(* Logix 5000 project; controller FV vendor 1 type 14 code 217 rev 31.11; software revision 31.00 *) (continued)
   FR_N10 : INT[265] := ([1] := 1, [2] := 4, [3] := 6, [6] := 6, [100] := 1, [101] := 2, [102] := 3, [103] := 3, [104] := 9, [105] := 9, [106] := 3, [200] := 2, [203] := 20, [204] := 191, [205] := 137, [206] := 100, [209] := 23, [215] := 14641, [216] := 11826, [217] := 13873, [218] := 11832, [219] := 12338, [220] := 13102, [221] := 49);   // FV_AGING Comms to FV Aging PL C
        [0]   // FV Unit Heartbeat
        [0].0   // FV_Aging PLC Heartbeat
        [100].0   // FV Routing (This)PLC Heartbeat
        [101]   // FV26 Routing Status to FV PLC
        [102]   // FV27 Routing Status to FV PLC
        [103]   // FV28 Routing Status to FV PLC
        [104]   // FV29 Routing Status to FV PLC
        [105]   // FV30 Routing Status to FV PLC
        [106]   // FV31 Routing Status to FV PLC
        [1]   // FV26 Aging Status from FV PLC
        [200].0   // FV_Aging_PLC Heartbeat Fault
        [200].1   // Enable Comms to FV Aging PLC
        [201]   // FV_Aging PLC Comms Control Block
        [2]   // FV27 Aging Status from FV PLC
        [3]   // FV28 Aging Status from FV PLC
        [4]   // FV29 Aging Status from FV PLC
        [5]   // FV30 Aging Status from FV PLC
        [6]   // FV31 Aging Status from FV PLC
   FR_N100 : INT[265] := ([2] := 1, [3] := 129, [6] := -1, [7] := -1, [8] := 2530, [9] := -1, [10] := 1, [15] := 1, [20] := -1, [21] := -1, [22] := -1, [23] := -1, [24] := -1, [25] := -1, [26] := -1, [30] := 226, [32] := 1000, [33] := 8, [35] := -1, [36] := -1, [40] := 26, [42] := 70, [47] := 50, [48] := 300, [49] := 32760, [57] := 2046, [70] := 32760, [71] := 32760, [72] := 32760, [73] := 32760, [74] := 32760, [75] := 32760, [100] := 22, [101] := 9, [102] := 14, [103] := 26, [104] := 25, [105] := 37, [106] := 28, [107] := 33, [108] := 41, [109] := 40, [110] := 74, [111] := 65, [112] := 70, [113] := 78, [114] := 77, [115] := -1, [116] := -1, [117] := -1, [118] := -1, [119] := -1, [120] := -1, [121] := -1, [122] := -1, [123] := -1, [124] := -1, [125] := -1, [126] := -1, [127] := -1,
        [128] := -1, [129] := -1, [130] := -1, [131] := -1, [132] := -1, [133] := -1, [134] := -1, [135] := -1, [136] := -1, [137] := -1, [138] := -1, [139] := -1, [140] := -1, [141] := -1, [142] := -1, [143] := -1, [144] := -1, [145] := -1, [146] := -1, [147] := -1, [148] := -1, [149] := -1);   // FV FILLING
        [0]   // FV_Fill Step
        [100]   // FV Filling Checklist Data
        [10]   // FV_Fill Idle Step Bits
        [10].0   // FV_Fill STEP Available
        [10].1   // FV_Fill STEP Clean
        [10].2   // FV_Fill STEP Command Data Check
        [10].3   // FV_Fill STEP Data in Limits Check
        [10].4   // FV_Fill STEP FV Vessel Status Check
        [10].6   // FV_Fill STEP Prestart Checks Failed
        [11]   // FV_Fill Running Step Bits
        [11].0   // FV_Fill STEP Initialise Transfer
        [11].1   // FV_Fill STEP Beer Chase
        [11].2   // FV_Fill STEP Valve Changeover
        [11].3   // FV_Fill STEP Filling
        [11].4   // FV_Fill Beer Transfer Complete
        [11].5   // FV_Fill Liquor Transfer Complete
        [11].8   // FV_Fill Step Transfer Complete
        [12]   // FV_Fill CIP Step Bits
        [12].0   // FV_Fill STEP CIP
        [12].1   // FV_Fill CIP Channel 1 Complete
        [12].2   // FV_Fill STEP Channel 2 CIP
        [12].3   // FV_Fill CIP Channel 2 Complete
        [13]   // FV_Fill Held Step Bits
        [13].1   // FV_Fill Faulted
        [14].0   // FV_Fill STEP Data in Limits Check Vessel Number OK
        [15].0   // FV_Fill Auto FV
        [16].2   // FV_Fill STEP Initialise Transfer All Systems at Prestart Failed
        [17].0   // MV_Fill Backup STEP Initialise Transfer
        [17].1   // FV_Fill Backup STEP Beer Chase
        [17].2   // FV_Fill Backup STEP Valve Changeover
        [17].3   // FV_Fill Backup STEP Filling
        [17].4   // FV_Fill Backup STEP Beer Transfer Complete
        [17].5   // FV_Fill Backup STEP Liquor Transfer Complete
        [17].6   // MV_Fill Backup STEP Flush to Drain
        [17].8   // FV_Fill Backup Step Transfer Complete
        [1]   // FV_Fill Backup Step
        [20]   // FV_Fill SCADA Download Vessel ID
        [21]   // FV_Fill SCADA Download Beer Chase Required
        [22]   // FV_Fill SCADA Download Fermenting Pressure
        [23]   // FV_Fill SCADA Download Chill Down Pressure
        [24]   // FV_Fill SCADA Download Chill Down Time
        [25]   // FV_Fill SCADA Download Chill Down Time
        [27]   // Final Gravity
        [2]   // FV_Fill Status
        [2].0   // FV_Fill STATUS Idle
        [2].1   // FV_Fill STATUS Running
        [2].2   // FV_Fill STATUS CIP
        [2].3   // FV_Fill STATUS Held
        [30]   // FV_Fill Vessel ID
        [31]   // FV_Fill Beer Chase Required
        [32]   // FV_Fill Fermenting Pressure
        [33]   // FV_Fill Chill Down Pressure
        [34]   // FV_Fill Chill Down Time
        [3]   // FV_Fill SCADA Prompts
        [3].0   // FV_Fill SCADA Prompts Start
        [3].1   // FV_Fill SCADA Prompts Hold
        [3].15   // FV_Fill SCADA Prompts Reset
        [3].2   // FV_Fill SCADA Prompts Continue
        [3].3   // FV_Fill SCADA Prompts Abort
        [3].4   // FV_Fill SCADA Prompts Cancel
        [3].5   // FV_Fill STEP SCADA Prompts Beer Transfer Complete
        [3].6   // FV_Fill STEP SCADA Prompts Liquor Transfer Complete
        [3].7   // FV_Fill SCADA Prompts Set for CIP
        [3].8   // FV_Fill SCADA Prompts Clear CIP Route
        [40]   // FV_Fill FV File Number
        [42]   // FV_Fill STEP Preset Chase Volume
        [43]   // FV_Fill STEP Actual Chase Pulses
        [44]   // FV_Fill STEP Actual Chase Volume
        [45]   // FV_Fill STEP Beer Tansfer Pulses
        [46]   // FV_Fill STEP Beer Tansfer Volume
        [47]   // Check Flow before Checking O2 Valve
        [49]   // Paraflow Totaliser
        [4]   // FV_Fill SCADA Commands
        [4].0   // FV_Fill SCADA Commands Start
        [4].4   // FV_Fill SCADA Commands Cancel
        [4].5   // FV_Fill STEP SCADA Commands Beer Transfer Complete
        [4].6   // FV_Fill STEP SCADA Commands Liquor Transfer Complete
        [4].7   // FV_Fill SCADA Commands Set for CIP
        [4].8   // FV_Fill SCADA Commands Clear CIP Route
        [50]   // FV_Fill Chase Countdown
        [57]   // FV_Fill Last Plant Fault
        [5]   // FV_Fill Last SCADA Commands
        [5].0   // FV_Fill SCADA Commands Start
        [60].0   // FV_Fill CIP Route Open
        [6]   // FV_Fill Plant Warning
        [70]   // FV26 Filling Totaliser
        [71]   // FV27 Filling Totaliser
        [72]   // FV28 Filling Totaliser
        [73]   // FV29 Filling Totaliser
        [74]   // FV30 Filling Totaliser
        [75]   // FV31 Filling Totaliser
        [7]   // FV_Fill Plant Fault
        [8]   // FV_Fill Log Message
        [9]   // FV_Fill Plant Item Fault
   FR_N100_6_alarm : ALARM_DIGITAL;
   FR_N100_6_Alarm_Ready : BOOL;
   FR_N100_6_Delayed : DINT := -1;
   FR_N100_6_Delayed_Timer : TIMER := (PRE := 1000);
   FR_N100_6_Fault_Returned : STRING;
   FR_N100_6_SQL_Done : DINT := -1;
   FR_N100_7_alarm : ALARM_DIGITAL;
   FR_N100_7_Alarm_Ready : BOOL;
   FR_N100_7_Delayed : DINT := -1;
   FR_N100_7_Delayed_Timer : TIMER := (PRE := 1000);
   FR_N100_7_Delayed_Timer2 : TIMER := (PRE := 1000);
   FR_N100_7_Fault_Returned : STRING;
   FR_N100_7_SQL_Done : DINT := -1;
   FR_N100_8_Delayed : DINT := 2530;
   FR_N100_8_Delayed_Timer : TIMER := (PRE := 1000);
   FR_N100_8_Event_Returned : STRING := 'FV26 FV Filling, Beer Fill Complete confirmed by Operator';
   FR_N100_8_SQL_Done : DINT;
   FR_N110 : INT[265] := ([2] := 1, [3] := 1, [6] := -1, [7] := -1, [8] := 2651, [9] := -1, [10] := 1, [15] := 1, [20] := -1, [21] := -1, [30] := 226, [40] := 26, [41] := 226, [50] := 511, [57] := 2015, [100] := 18, [101] := 20, [102] := 23, [103] := 10, [104] := 15, [105] := 38, [106] := 29, [107] := 34, [108] := 75, [109] := 66, [110] := 71, [111] := 2, [112] := -1, [113] := -1, [114] := -1, [115] := -1, [116] := -1, [117] := -1, [118] := -1, [119] := -1, [120] := -1, [121] := -1, [122] := -1, [123] := -1, [124] := -1, [125] := -1, [126] := -1, [127] := -1, [128] := -1, [129] := -1, [130] := -1, [131] := -1, [132] := -1, [133] := -1, [134] := -1, [135] := -1, [136] := -1, [137] := -1, [138] := -1, [139] := -1, [140] := -1, [141] := -1, [142] := -1, [143] := -1, [144] := -1,
        [145] := -1, [146] := -1, [147] := -1, [148] := -1, [149] := -1);   // GREEN BEER Green Beer Main
        [0]   // Green Beer STEP
        [100]   // Green Beer Checklist Data
        [10]   // Green Beer Idle Bits
        [10].0   // Green Beer Step Bits Idle
        [10].1   // Green Beer Step Bits Clean
        [10].2   // Green Beer Wait for SCADA Data
        [10].3   // Green Beer Check SCADA Data
        [10].4   // Green Beer Check Vessel Status
        [10].5   // FV>MV STEP Prestart Check
        [11]   // Green Beer Running Bits
        [11].0   // Green Beer STEP Initialise
        [11].1   // FV>MV STEP Open Drain
        [11].2   // FV>MV STEP Beer Chase
        [11].3   // Green Beer STEP Beer Transfer
        [11].4   // Green Beer FV Volume Transferred or Empty
        [11].5   // Green Beer STEP Water Chase
        [11].6   // FV>MV STEP Water Flush Complete
        [11].7   // FV>MV STEP Manual Transfer
        [11].8   // Green Beer STEP Transfer Complete
        [12]   // Green Beer CIP Bits
        [12].0   // FV26-31 Green Beer Main Channel 1 CIP
        [12].1   // Green Beer Channel 1 CIP Complete
        [12].2   // FV26-31 Green Beer Main Channel 2 CIP
        [12].3   // Green Beer Channel 2 CIP Complete
        [12].4   // FV26-31 Green Beer Main Channel 1 CIP
        [12].5   // FV26-31 Green Beer Main Channel 1 CIP Complete
        [12].6   // FV26-31 Green Beer Main Channel 2 CIP
        [12].7   // FV26-31 Green Beer Main Channel 2 CIP Complete
        [13]   // Green Beer Hold Bits
        [13].0   // Green Beer Transfer Held
        [13].1   // Green Beer Transfer Faulted
        [14].0   // Green Beer Auto FV
        [15]   // FV>MV Flags
        [15].0   // Green Beer FV Vessel is Auto
        [15].1   // FV>MV STEP Prestart Check OK
        [15].2   // FV>MV Prestart Check Failed
        [15].3   // FV>MV Beer Available
        [15].4   // FV>MV Volume Transferred
        [15].5   // FV>MV Chase Water Open
        [15].6   // FV>MV Chase Water Closed
        [15].7   // FV>MV FV Empty
        [18].0   // Green Beer Extended
        [1]   // Green Beer Backup Step
        [20]   // Green Beer Vessel ID
        [21]   // Green Beer Volume to Transfer
        [22]   // FV>MV_ Volume to Transfer
        [23]   // Vessel Initial Volume
        [24]   // Vessel Transferred Volume
        [2].0   // Green Beer Idle
        [2].1   // Green Beer Running
        [2].2   // Green Beer CIP
        [2].3   // Green Beer Held
        [31]   // Green Beer Transfer Target
        [3].0   // Green Beer PROMPTS Start
        [3].1   // Green Beer SCADA Prompt Hold
        [3].15   // Green Beer SCADA Prompt Reset
        [3].2   // Green Beer SCADA Prompt Continue
        [3].3   // Green Beer SCADA Prompt Abort
        [3].4   // Green Beer PROMPTS Cancel
        [3].5   // Green Beer STEP SCADA Prompts Beer Transfer Complete
        [3].6   // Green Beer STEP SCADA Prompts Extend Transfer
        [3].7   // Green Beer STEP SCADA Prompts Flush Main
        [3].8   // Green Beer STEP SCADA Prompts End Transfer
        [3].9   // Green Beer STEP SCADA Prompts End Flush
        [40]   // Green Beer Vessel File Number
        [4]   // Green Beer SCADA Command
        [4].0   // Green Beer COMMANDS Start
        [4].1   // Green Beer SCADA Command Hold
        [4].15   // Green Beer SCADA Command Reset
        [4].2   // Green Beer SCADA Command Continue
        [4].3   // Green Beer SCADA Command Abort
        [4].4   // Green Beer COMMANDS Cancel
        [4].5   // Green Beer STEP SCADA Commands Beer Transfer Complete
        [4].6   // Green Beer STEP SCADA Command Extend Transfer
        [4].7   // Green Beer STEP SCADA Commands Flush Main
        [4].8   // Green Beer STEP SCADA Commands End Transfer
        [4].9   // Green Beer STEP SCADA Commands End Flush
        [50]   // Vessel Initial Volume
        [51]   // Green Beer Volume Transferred
        [52]   // Green Beer Volume Remaining
        [57]   // Green Beer Last Plant Fault
        [5]   // Green Beer Last SCADA Command
        [60].0   // FV26-31 Green Beer Main CIP Route Open
        [6]   // Green Beer Warning
        [7]   // Green Beer Faults
        [8]   // Green Beer Log Message
        [9]   // FV26-31 Green Beer Main Plant Item Fault
   FR_N110_6_alarm : ALARM_DIGITAL;
   FR_N110_6_Alarm_Ready : BOOL;
   FR_N110_6_Delayed : DINT := -1;
   FR_N110_6_Delayed_Timer : TIMER := (PRE := 1000);
   FR_N110_6_Fault_Returned : STRING;
   FR_N110_6_SQL_Done : DINT := -1;
   FR_N110_7_alarm : ALARM_DIGITAL;
   FR_N110_7_Alarm_Ready : BOOL;
   FR_N110_7_Delayed : DINT := -1;
   FR_N110_7_Delayed_Timer : TIMER := (PRE := 1000);
   FR_N110_7_Delayed_Timer2 : TIMER := (PRE := 1000);
   FR_N110_7_Fault_Returned : STRING;
   FR_N110_7_SQL_Done : DINT := -1;
   FR_N110_8_Delayed : DINT := 2651;
   FR_N110_8_Delayed_Timer : TIMER := (PRE := 1000);
   FR_N110_8_Event_Returned : STRING := 'FV26 FV26-31 green beer main CIP completed.';
   FR_N110_8_SQL_Done : DINT;
   FR_N120 : INT[265] := ([2] := 1, [3] := 1, [6] := -1, [7] := -1, [8] := 2721, [9] := -1, [10] := 1, [15] := 2, [20] := -1, [21] := -1, [22] := -1, [23] := -1, [24] := -1, [25] := -1, [26] := -1, [29] := 227, [30] := 8, [31] := 200, [32] := 300, [33] := 60, [34] := 120, [35] := 1200, [36] := 35, [40] := 26, [42] := 99, [47] := 2011, [50] := 100, [51] := 500, [52] := 2, [53] := 10, [55] := 2, [56] := 100, [57] := 100, [58] := 5, [100] := 19, [101] := 21, [102] := 24, [103] := 11, [104] := 16, [105] := 39, [106] := 30, [107] := 35, [108] := 76, [109] := 67, [110] := 72, [111] := 1, [112] := -1, [113] := -1, [114] := -1, [115] := -1, [116] := -1, [117] := -1, [118] := -1, [119] := -1, [120] := -1, [121] := -1, [122] := -1, [123] := -1, [124] := -1, [125] := -1,
        [126] := -1, [127] := -1, [128] := -1, [129] := -1, [130] := -1, [131] := -1, [132] := -1, [133] := -1, [134] := -1, [135] := -1, [136] := -1, [137] := -1, [138] := -1, [139] := -1, [140] := -1, [141] := -1, [142] := -1, [143] := -1, [144] := -1, [145] := -1, [146] := -1, [147] := -1, [148] := -1, [149] := -1);   // YEAST CROP Yeast Cropping Main
        [0]   // Yeast Cropping Step
        [100]   // Yeast Cropping Checklist Data
        [10]   // Yeast Cropping Idle Step Bits
        [10].0   // Yeast Removal STEP Available
        [10].1   // Yeast Removal STEP Clean
        [10].2   // Yeast Removal STEP Command Data Check
        [10].3   // Yeast Removal STEP Data in Limits Check
        [10].4   // Yeast Removal STEP FV Vessel Status Check
        [11]   // Yeast Cropping Running Step Bits
        [11].0   // Yeast Cropping STEP Initialise Transfer
        [11].1   // Yeast Cropping STEP Open Route
        [11].2   // Yeast Cropping STEP Minimum Speed
        [11].3   // Yeast Cropping Step Ramp Up
        [11].4   // Yeast Cropping STEP Maximum Speed
        [11].5   // Yeast Cropping Done
        [11].6   // Yeast Cropping Flush
        [11].8   // Yeast Cropping Complete
        [12]   // Yeast Cropping CIP Step Bits
        [12].0   // Yeast Removal Channel 1 CIP
        [12].1   // Yeast Removal Channel 1 CIP Complete
        [12].2   // Yeast Removal Channel 2 CIP
        [12].3   // Yeast Removal Channel 2 CIP Complete
        [13]   // Yeast Cropping Held Step Bits
        [13].1   // Yeast Cropping Fault
        [14].0   // Yeast Removal STEP Data in Limits Check Vessel Number OK
        [15].0   // Yeast Removal Auto FV Pump1
        [15].1   // Yeast Removal Pump2
        [15].2   // Yeast Removal Pump3
        [16].0   // FV26-31 Channel 1 CIP Reset Complete Flag
        [16].1   // FV1-17 Channel 1 CIP Reset Complete Flag
        [16].2   // FV18-25 Channel 1 CIP Reset Complete Flag
        [16].3   // FV26-31 Channel 2 CIP Reset Complete Flag
        [16].4   // FV1-17 Channel 2 CIP Reset Complete Flag
        [16].5   // FV18-25 Channel 2 CIP Reset Complete Flag
        [16].6   // Yeast Removal Pump3 CIP Ch2 Selected
        [17].0   // FV26-31 Channel 1 CIP OSR to reset Complete Flag
        [17].1   // FV1-17 Channel 1 CIP OSR to reset Complete Flag
        [17].2   // FV18-25 Channel 1 CIP OSR to reset Complete Flag
        [17].3   // FV26-31 Channel 2 CIP OSR to reset Complete Flag
        [17].4   // FV1-17 Channel 2 CIP OSR to reset Complete Flag
        [17].5   // FV18-25 Channel 2 CIP OSR to reset Complete Flag
        [1]   // Yeast Cropping Backup Step
        [20]   // Yeast Cropping SCADA Download Vessel ID
        [21]   // Yeast Cropping SCADA Download Minimum Speed
        [22]   // Yeast Cropping SCADA Download Maximum Speed
        [23]   // Yeast Cropping SCADA Download Minimum Speed Duration
        [24]   // Yeast Cropping SCADA Download Ramp Up Duration
        [25]   // Yeast Cropping SCADA Download Maximum Speed Duration
        [26]   // Yeast Cropping SCADA Download Flush Duration
        [2]   // Yeast Cropping Status
        [2].0   // Yeast Removal Status Idle
        [2].1   // Yeast Removal Status Running
        [2].2   // Yeast Removal Status CIP
        [2].3   // Yeast Removal Status Held
        [30]   // Yeast Cropping Vessel ID
        [31]   // Yeast Cropping Minimum Speed
        [32]   // Yeast Cropping Maximum Speed
        [33]   // Yeast Cropping Minimum Speed Duration
        [34]   // Yeast Cropping Ramp Up Duration
        [35]   // Yeast Cropping Maximum Speed Duration
        [36]   // Yeast Cropping Flush Duration
        [3]   // Yeast Cropping SCADA Prompts
        [3].0   // Yeast Removal SCADA Prompts Start
        [3].1   // Yeast Removal SCADA Prompts Hold
        [3].15   // Yeast Removal SCADA Prompts Reset
        [3].2   // Yeast Removal SCADA Prompts Continue
        [3].3   // Yeast Removal SCADA Prompts Abort
        [3].4   // Yeast Removal SCADA Prompts Cancel
        [3].5   // Yeast Removal SCADA Prompts Flush
        [3].6   // Yeast Removal SCADA Prompts Complete
        [40]   // Yeast Cropping FV File Number
        [41]   // Yeast Cropping Pump Speed
        [42]   // Ramp Up Current Time
        [47]   // Yeast Cropping Last Plant Fault
        [4]   // Yeast Cropping SCADA Commands
        [4].0   // Yeast Removal SCADA Commands Start
        [4].1   // Yeast Removal SCADA Commands Hold
        [4].2   // Yeast Removal SCADA Commands Continue
        [4].3   // Yeast Removal SCADA Commands Abort
        [4].4   // Yeast Removal SCADA Commands Cancel
        [4].5   // Yeast Removal SCADA Commands Flush
        [4].6   // Yeast Removal SCADA Commands Complete
        [58]   // Yeast Removal Flush Duration
        [5]   // Yeast Cropping Last SCADA Commands
        [60].0   // FV26-31 Yeast Main CIP Route Open
        [62]   // Yeast Cropping Step Time Remaining
        [6]   // Yeast Cropping Plant Warning
        [7]   // Yeast Cropping Plant Fault
        [8]   // Yeast Cropping Log Message
        [9]   // Yeast Cropping Plant Item Fault
   FR_N120_17_0_Storagebit : BOOL;
   FR_N120_17_1_Storagebit : BOOL;
   FR_N120_17_2_Storagebit : BOOL;
   FR_N120_17_3_Storagebit : BOOL;
   FR_N120_17_4_Storagebit : BOOL;
   FR_N120_17_5_Storagebit : BOOL;
   FR_N120_6_alarm : ALARM_DIGITAL;
   FR_N120_6_Alarm_Ready : BOOL;
   FR_N120_6_Delayed : DINT := -1;
   FR_N120_6_Delayed_Timer : TIMER := (PRE := 1000);
   FR_N120_6_Fault_Returned : STRING;
   FR_N120_6_SQL_Done : DINT := -1;
   FR_N120_7_alarm : ALARM_DIGITAL;
   FR_N120_7_Alarm_Ready : BOOL;
   FR_N120_7_Delayed : DINT := -1;
   FR_N120_7_Delayed_Timer : TIMER := (PRE := 1000);
   FR_N120_7_Delayed_Timer2 : TIMER := (PRE := 1000);
   FR_N120_7_Fault_Returned : STRING;
   FR_N120_7_SQL_Done : DINT := -1;
   FR_N120_8_Delayed : DINT := 2721;
   FR_N120_8_Delayed_Timer : TIMER := (PRE := 1000);
   FR_N120_8_Event_Returned : STRING := 'FV8 Yeast Cropping, Complete confirmed by Operator';
   FR_N120_8_SQL_Done : DINT;
   FR_N13 : INT[265] := ([2] := 1, [3] := 1, [6] := 2, [103] := 226, [104] := -1, [105] := 1, [108] := 1, [200] := 2, [201] := 4312, [203] := 20, [204] := 12, [205] := 137, [206] := 100, [209] := 23, [215] := 14641, [216] := 11826, [217] := 13873, [218] := 11832, [219] := 12338, [220] := 13102, [221] := 52);   // MV_ROUTE Comms to MV Routing PLC
        [0].0   // MV_Routing_Unit Heartbeat
        [100].0   // FV_Routing(This PLC) Heartbeat
        [101]   // MV_Routing_Unit_PLC_ Echo of MV>FV Transfer Step
        [102]   // MV_Routing_Unit_PLC_ Echo of FV Vessel
        [103]   // MV_Routing_Unit_PLC_ Echo of Vessel ID
        [104]   // MV_Routing_Unit_PLC_ Plant Item Fault
        [105]   // FV>MV Flags
        [105].3   // FV>MV Beer Available
        [106]   // Centrifuge 1 Pulse Count
        [107]   // Centrifuge 2 Pulse Count
        [108].0   // Green Beer Main Ready for centrifuge
        [108].1   // FV26 Ready for centrifuge
        [108].2   // FV27 Ready for centrifuge
        [108].3   // FV28 Ready for centrifuge
        [108].4   // FV29 Ready for centrifuge
        [108].5   // FV30 Ready for centrifuge
        [108].6   // FV31 Ready for centrifuge
        [1]   // MV_Routing_Unit_PLC_ MV>FV Transfer Step
        [200].0   // MV_Routing_Unit Heartbeat Fault
        [200].1   // Enable Comms to MV Routing Unit
        [201]   // MV_Routing_Unit Comms Control Block
        [2]   // MVFV_CIP_Unit_PLC Status
        [3]   // MV_Routing_Unit_PLC_ FV to Transfer
        [4]   // MV_Routing_Unit_PLC_ Volume to Transfer
        [5].0   // Auto MV Filling at High Level
        [6].0   // Count Centrifuge Pulses
        [6].1   // Clear Centrifuge Pulse Counts
   FR_N130 : INT[265] := ([2] := 1, [3] := 1, [6] := -1, [7] := 2833, [8] := 2850, [9] := 2060, [10] := 1, [15] := 1, [20] := -1, [21] := -1, [22] := -1, [23] := -1, [24] := -1, [25] := -1, [26] := -1, [30] := 229, [32] := -1, [33] := -1, [34] := -1, [35] := -1, [36] := -1, [40] := 29, [47] := 2057, [61] := 3, [62] := 4, [100] := 57, [101] := 62, [102] := 59, [103] := 58, [104] := 79, [105] := 56, [106] := 55, [107] := 54, [108] := 60, [109] := 5, [110] := -1, [111] := -1, [112] := -1, [113] := -1, [114] := -1, [115] := -1, [116] := -1, [117] := -1, [118] := -1, [119] := -1, [120] := -1, [121] := -1, [122] := -1, [123] := -1, [124] := -1, [125] := -1, [126] := -1, [127] := -1, [128] := -1, [129] := -1, [130] := -1, [131] := -1, [132] := -1, [133] := -1, [134] := -1,
        [135] := -1, [136] := -1, [137] := -1, [138] := -1, [139] := -1, [140] := -1, [141] := -1, [142] := -1, [143] := -1, [144] := -1, [145] := -1, [146] := -1, [147] := -1, [148] := -1, [149] := -1);   // FILTRATE Filtrate Return
        [0]   // Filtrate Return Step
        [100]   // Filtrate Return Checklist Data
        [10]   // Filtrate Return Idle Step Bits
        [10].0   // Filtrate Return STEP Available
        [10].1   // Filtrate Return STEP Clean
        [10].2   // Filtrate Return STEP Command Data Check
        [10].3   // Filtrate Return STEP Data in Limits Check
        [10].4   // Filtrate Return STEP FV Vessel Status Check
        [11]   // Filtrate Return Running Step Bits
        [11].0   // Filtrate Return STEP Initialise Transfer
        [11].1   // Filtrate Return STEP Open Route
        [11].2   // Filtrate Return STEP Drain Gas Main
        [11].3   // Filtrate Return Step Drain the Mains First
        [11].4   // Filtrate Return STEP Maximum Speed
        [11].5   // Filtrate Return STEP Flush
        [12]   // Filtrate Return CIP Step Bits
        [12].0   // Filtrate Return Channel 1 CIP
        [12].1   // Filtrate Return Channel 1 CIP Complete
        [12].2   // Filtrate Return Channel 2 CIP
        [12].3   // Filtrate Return Channel 2 CIP Complete
        [12].4   // Filtrate Return FRV1 Ch1 CIP
        [12].5   // Filtrate Return FRV1 Ch1 CIP Complete
        [12].6   // Filtrate Return FRV1 Ch2 CIP
        [12].7   // Filtrate Return FRV1 Ch2 CIP Complete
        [13]   // Filtrate Return Held Step Bits
        [13].1   // Filtrate Return Fault
        [14].0   // Filtrate Return STEP Data in Limits Check Vessel Number OK
        [15].0   // Filtrate Return Auto FV
        [1]   // Filtrate Return Backup Step
        [20]   // Filtrate Return SCADA Download Vessel ID
        [2]   // Filtrate Return Status
        [2].0   // Filtrate Return Status Idle
        [2].1   // Filtrate Return Status Running
        [2].2   // Filtrate Return Status CIP
        [2].3   // Filtrate Return Status Held
        [30]   // Filtrate Return Vessel ID
        [31]   // Filtrate Return Drain the Mains First
        [3]   // Filtrate Return SCADA Prompts
        [3].0   // Filtrate Return SCADA Prompts Start
        [3].1   // Filtrate Return SCADA Prompts Hold
        [3].15   // Filtrate Return SCADA Prompts Reset
        [3].2   // Filtrate Return SCADA Prompts Continue
        [3].3   // Filtrate Return SCADA Prompts Abort
        [3].4   // Filtrate Return SCADA Prompts Cancel
        [3].5   // Filtrate Return SCADA Prompt Filtrate Return Complete
        [40]   // Filtrate Return FV File Number
        [41]   // Minimum Speed
        [47]   // Filtrate Return Last Plant Fault
        [4]   // Filtrate Return SCADA Commands
        [4].5   // Filtrate Return SCADA Command Filtrate Return Complete
        [50]   // Filtrate Return Minimum Speed
        [51]   // Filtrate Return Maximum Speed
        [52]   // Filtrate Return Minimum Speed Duration
        [53]   // Filtrate Return Ramp Duration
        [54]   // Filtrate Return Ramp Current Time
        [55]   // Filtrate Return Maximum Speed Duration
        [56]   // Filtrate Return Ramp Speed
        [57]   // Filtrate Return Pump Speed
        [58]   // Filtrate Return Flush Duration
        [5]   // Filtrate Return Last SCADA Commands
        [60].0   // FV26-31 Filtrate Main CIP Route Open
        [61]   // Filtrate Tank Mode
        [62].0   // Filtrate Tank Process
        [62].1   // Filtrate Tank Tank CIP
        [62].2   // Filtrate Tank Line CIP
        [63].0   // FRV1 Request Channel 1 CIP
        [63].1   // FRV1 Request Channel 2 CIP
        [6]   // Filtrate Return Plant Warning
        [7]   // Filtrate Return Plant Fault
        [8]   // Filtrate Return Log Message
        [9]   // Filtrate Return Plant Item Fault
   FR_N130_6_alarm : ALARM_DIGITAL;
   FR_N130_6_Alarm_Ready : BOOL;
   FR_N130_6_Delayed : DINT := -1;
   FR_N130_6_Delayed_Timer : TIMER := (PRE := 1000);
   FR_N130_6_Fault_Returned : STRING;
   FR_N130_6_SQL_Done : DINT := -1;
   FR_N130_7_alarm : ALARM_DIGITAL;
   FR_N130_7_Alarm_Ready : BOOL := 1;
   FR_N130_7_Delayed : DINT := 2833;
   FR_N130_7_Delayed_Timer : TIMER := (PRE := 1000);
   FR_N130_7_Delayed_Timer2 : TIMER := (PRE := 1000);
   FR_N130_7_Fault_Returned : STRING := 'FV29 Filtrate Return, Filtrate Tank not set to Line CIP.';
   FR_N130_7_SQL_Done : DINT := -1;
   FR_N130_8_Delayed : DINT := 2850;
   FR_N130_8_Delayed_Timer : TIMER := (PRE := 1000);
   FR_N130_8_Event_Returned : STRING := 'FV29 Filtrate Return Main, CIP aborted.';
   FR_N130_8_SQL_Done : DINT;
   FR_N14 : INT[265] := ([11] := 1, [12] := 1, [13] := 8, [101] := 24, [102] := 7, [103] := -1, [104] := 2000, [109] := 5, [110] := 4, [111] := 24, [112] := 7, [113] := -1, [114] := -4, [200] := 2, [201] := 8192, [203] := 20, [204] := 112, [205] := 137, [206] := 100, [209] := 23, [215] := 14641, [216] := 11826, [217] := 13873, [218] := 11832, [219] := 12338, [220] := 13102, [221] := 54);   // MVFV CIP Comms to MVFV CIP Un it PLC
        [0].0   // MVFV CIP PLC Heartbeat
        [101]   // CIP Available for Ch1 CIP Flags
        [101].0   // FV26 Available for Ch1 CIP
        [101].1   // FV27 Available for Ch1 CIP
        [101].2   // FV28 Available for Ch1 CIP
        [101].3   // FV29 Available for Ch1 CIP
        [101].4   // FV30 Available for Ch1 CIP
        [101].5   // FV31 Available for Ch1 CIP
        [101].6   // Filtrate Tank Available for CIP
        [102].0   // FV26-31 Green Beer Main Available for Ch1 CIP
        [102].1   // FV26-31 Yeast Cropping Main Available for Ch1 CIP
        [102].2   // FV26-31 Filtrate Return Main Available for Ch1 CIP
        [103]   // Channel 1 CIP Fault
        [104]   // Channel 1 CIP Status
        [104].0   // Channel 1 CIP Route Open
        [104].1   // Channel 1 CIP Complete
        [110].0   // Copy FV1-17 Yeast Pump 2 CIP Return Proxy to MVFV CIP Unit
        [110].1   // Copy FV18-25 Yeast Pump 3 CIP Return Proxy to MVFV CIP Unit
        [110].2   // Copy FV26-31 Yeast Pump 1 CIP Return Proxy to MVFV CIP Unit
        [111]   // CIP Available for Ch2 CIP Flags
        [113]   // Channel 2 CIP Fault
        [114]   // Channel 2 CIP Status
        [114].0   // Channel 2 CIP Route Open
        [114].1   // Channel 2 CIP Complete
        [11]   // CIP Channel 2 Route
        [12]   // CIP Channel 2 Program
        [13]   // CIP Channel 2 Vessel
        [14].0   // CIP Channel 2 Active
        [14].1   // CIP Channel 2 Open Route
        [14].2   // CIP Channel 2 Run Return Pump
        [14].3   // CIP Channel 2 Complete
        [14].4   // Vessel Status Channel 2 CIP Acknowledge Alarm
        [14].5   // CIP Channel 2 Detergent Circulating
        [14].6   // CIP Channel 2 Flow Established
        [1]   // CIP Channel 1 Route
        [200].0   // MVFV CIP PLC Heartbeat Fault
        [200].1   // Enable Comms to MVFV CIP Unit PLC
        [201]   // Comms to MVFV CIP Unit PLC
        [2]   // CIP Channel 1 Program
        [3]   // CIP Channel 1 Vessel
        [4].0   // CIP Channel 1 Active
        [4].1   // CIP Channel 1 Open Route
        [4].2   // CIP Channel 1 Run Return Pump
        [4].3   // CIP Channel 1 Complete
        [4].4   // Vessel Status Channel 1 CIP Acknowledge Alarm
        [4].5   // CIP Channel 1 Detergent Circulating
        [4].6   // CIP Channel 1 Flow Established
   FR_N140 : INT[265] := ([1] := 1, [3] := 2060);   // CIP
        [0].0   // FV26-31 Filling Main Request Channel 1 CIP
        [0].1   // FV26-31 Green Beer Main Request Channel 1 CIP
        [0].2   // FV26-31 Yeast Main Request Channel 1 CIP
        [0].3   // FV26-31 Filtrate Main Request Channel 1 CIP
        [0].4   // FV1-17 Yeast Main Request Channel 1 CIP
        [0].5   // FV18-25 Yeast Main Request Channel 1 CIP
        [0].6   // FRV1 Request Channel 1 CIP
        [10].0   // FV26-31 Filling Main Request Channel 2 CIP
        [10].1   // FV26-31 Green Beer Main Request Channel 2 CIP
        [10].2   // FV26-31 Yeast Main Request Channel 2 CIP
        [10].3   // FV26-31 Filtrate Main Request Channel 2 CIP
        [10].4   // FV1-17 Yeast Main Request Channel 2 CIP
        [10].5   // FV18-25 Yeast Main Request Channel 2 CIP
        [10].6   // FRV1 Request Channel 2 CIP
        [13]   // MV_Mains_CIP-Ch2 Plant Item Fault
        [1].0   // Do NOT Control Return Pump on Vessel Low Level
        [20].0   // Any Vessel on CIP
        [3]   // FV_Mains_CIP-Ch1 Plant Item Fault
   FR_N142 : INT[265];   // CIP
        [1]   // FV_Mains_CIP Selected Main
   FR_N143 : INT[265];   // CIP
   FR_N150 : INT[265];   // Original N File From SLC, No Description Available
        [14].0   // FV_Vessel_CIP Selected Vessel Valid Number
        [6].1   // FV_Routing(This PLC) Channel 1 Active
   FR_N160 : INT[265] := ([0] := 231, [1] := 3, [3] := 4, [5] := 6, [6] := 8, [7] := -1, [8] := 13231, [9] := -1, [10] := 1143, [11] := 8392, [12] := 1600, [13] := 2715, [14] := 529, [15] := 1144, [16] := 789, [17] := 8043, [18] := 32, [19] := 7794, [21] := 17, [22] := -125, [23] := 50, [24] := -75, [25] := -175, [26] := 1000, [27] := 8, [29] := 10, [30] := 21, [33] := 1, [37] := 600, [38] := 1144, [52] := 1, [60] := 16, [68] := 5323, [69] := 172, [100] := 42, [101] := 48, [102] := 54, [103] := 8, [104] := 88, [105] := 9, [106] := 10, [107] := 11, [108] := 12, [109] := -1, [110] := -1, [111] := -1, [112] := -1, [113] := -1, [114] := -1, [115] := -1, [116] := -1, [117] := -1, [118] := -1, [119] := -1, [120] := -1, [121] := -1, [122] := -1, [123] := -1, [124] := -1, [125] := -1,
        [126] := -1, [127] := -1, [128] := -1, [129] := -1, [130] := -1, [131] := -1, [132] := -1, [133] := -1, [134] := -1, [135] := -1, [136] := -1, [137] := -1, [138] := -1, [139] := -1, [140] := -1, [141] := -1, [142] := -1, [143] := -1, [144] := -1, [145] := -1, [146] := -1, [147] := -1, [148] := -1, [149] := -1, [200] := 120, [201] := 160);   // VESSEL Vessel Working Direc tory
        [0]   // Vessel ID
        [10]   // Vessel Level
        [11]   // Vessel Damped Level
        [12]   // Radius of Cone (mm)
        [13]   // Height of Cone (mm)
        [14]   // Vessel Volume (HL)
        [15]   // Pressure Difference Bottom - Top - Calibration (psi)
        [16]   // Pressure Difference Bottom - Top - Calibration (bar)
        [17]   // Height of column of water
        [18]   // Brewers Gravity
        [19]   // Height of column of beer
        [1]   // Vessel Status 0=Clean,1=Fill,2=Par t,3=Ferment,4=?,5=?, 6=?,7=?,8=Emptying,9 =Dirty,10-13=CIP
        [200]   // Checklist File Number
        [20]   // Vessel Step Bits
        [20].0   // Vessel Status Idle
        [20].1   // Vessel Status Top Pressure
        [20].2   // Vessel Status Chill Down
        [20].3   // Vessel Status Vent
        [20].5   // Vessel Status Channel 1 CIP
        [20].6   // Vessel Status Channel 1 CIP Complete
        [20].7   // Vessel Status Channel 2 CIP
        [20].8   // Vessel Status Channel 2 CIP Complete
        [21]   // Vessel Step Flags
        [21].0   // Vessel Top Pressure Control Over Pressure
        [21].1   // Vessel Top Pressure Control Under Pressure
        [21].12   // Vessel CIP Drain Down
        [21].2   // Vessel Top Pressure Control Zero Crossing
        [21].4   // Vessel Top Pressure Control Open Vent
        [21].5   // Vessel Top Pressure Control Open Vent Actuator
        [21].6   // Over Top Pressure Limit
        [22]   // Vessel Top Pressure Control Setpoint
        [23]   // Vessel Top Pressure Control Deadband
        [24]   // Vessel Top Pressure Control Upper Limit
        [25]   // Vessel Top Pressure Control Lower Limit
        [29]   // Vessel Top Pressure Chill Down Current Time
        [2]   // Vessel Level Probes
        [2].0   // FV Vessel High Level Probe
        [2].1   // FV Vessel Low Level Probe
        [30]   // Vessel Status Time since Clean
        [32]   // Vessel CIP Selected
        [32].0   // Channel 1 CIP Request
        [32].1   // Channel 2 CIP Request
        [33].1   // Vessel Rotocheck Fault
        [38]   // Vessel Pressure Difference Bottom-Top (psi)
        [39]   // Vessel Pressure Difference Calibration Offset
        [3]   // Top Pressure Status 0=Idle,1=Fill,2=Top Pressure,3=Chill Down,4=Vent,5=Emptyi ng,6=Ready for CIP
        [40]   // Yeast CroppingStatus 0=Not Done 1=Running 2=Done 3=Done+48hrs
        [41]   // Yeast Cropping Started Tally
        [42]   // Yeast Cropping Completed Tally
        [43]   // Vessel Hours since Yeast Cropping
        [4]   // Vessel Yeast Status
        [4].1   // Vessel Yeast Status Filtrate Return
        [50]   // Vessel Filtrate Status 0=Not Done 1=Running 2=Done
        [51]   // Vessel Filtrate Tally
        [52].0   // Vessel Filtrate Returning
        [52].1   // Vessel Filtrate Drain Back
        [5]   // Vessel Aging Status 1=Rise,2=Top, 3=Reduce,4=Hold, 5=Chill Down,6=Final
        [60].0   // Top Pressure Status Idle
        [60].1   // Top Pressure Status Filling
        [60].2   // Top Pressure Status Top Pressure
        [60].3   // Top Pressure Status Chill Down
        [60].4   // Top Pressure Status Vent
        [60].5   // Top Pressure Status Emptying
        [60].6   // Top Pressure Status Ready for CIP
        [68]   // Vessel Volume from paraflow
        [6]   // Vessel Valve Routes
        [7]   // Vessel Top Pressure Control Actual Pressure
        [8]   // Vessel Log Message
        [9]   // Vessel Item Fault
   FR_N170 : INT[265] := ([2] := 1, [3] := 1, [10] := 1, [100] := 3, [101] := -1, [102] := -1, [103] := -1, [104] := -1, [105] := -1, [106] := -1, [107] := -1, [108] := -1, [109] := -1, [110] := -1, [111] := -1, [112] := -1, [113] := -1, [114] := -1, [115] := -1, [116] := -1, [117] := -1, [118] := -1, [119] := -1, [120] := -1, [121] := -1, [122] := -1, [123] := -1, [124] := -1, [125] := -1, [126] := -1, [127] := -1, [128] := -1, [129] := -1, [130] := -1, [131] := -1, [132] := -1, [133] := -1, [134] := -1, [135] := -1, [136] := -1, [137] := -1, [138] := -1, [139] := -1, [140] := -1, [141] := -1, [142] := -1, [143] := -1, [144] := -1, [145] := -1, [146] := -1, [147] := -1, [148] := -1, [149] := -1);   // Original N File From SLC, No Description Available
        [0]   // Yeast Cropping FV1-17 Step
        [10]   // Yeast Cropping FV1-17 Idle Step Bits
        [10].0   // Yeast Cropping FV1-17 Available
        [10].1   // Yeast Cropping FV1-17 Clean
        [10].2   // Yeast Cropping FV1-17 Command Data Check
        [10].3   // Yeast Cropping FV1-17 Data in Limits Check
        [10].4   // Yeast Cropping FV1-17 FV Vessel Status Check
        [11]   // Yeast Cropping FV1-17 Running Step Bits
        [11].0   // Yeast Cropping FV1-17 Initialise Transfer
        [11].1   // Yeast Cropping FV1-17 Open Route
        [11].2   // Yeast Cropping FV1-17 Minimum Speed
        [11].3   // Yeast Cropping FV1-17 Ramp Up
        [11].4   // Yeast Cropping FV1-17 Maximum Speed
        [11].5   // Yeast Cropping FV1-17 Done
        [11].6   // Yeast Cropping FV1-17 Flush
        [12]   // Yeast Cropping FV1-17 CIP Step Bits
        [12].0   // Yeast Cropping FV1-17 Channel 1 CIP
        [12].1   // Yeast Cropping FV1-17 Channel 1 CIP Complete
        [12].2   // Yeast Cropping FV1-17 Channel 2 CIP
        [12].3   // Yeast Cropping FV1-17 Channel 2 CIP Complete
        [13]   // Yeast Cropping FV1-17 Held Step Bits
        [14].0   // Yeast Cropping FV1-17 Data in Limits Check Vessel Number OK
        [15].0   // Yeast Cropping FV1-17 Auto FV
        [1]   // Yeast Cropping FV1-17 Backup Step
        [20]   // Yeast Cropping FV1-17 SCADA Download Vessel ID
        [21]   // Yeast Cropping FV1-17 SCADA Download Minimum Speed
        [22]   // Yeast Cropping FV1-17 SCADA Download Maximum Speed
        [23]   // Yeast Cropping FV1-17 SCADA Download Minimum Speed Duration
        [24]   // Yeast Cropping FV1-17 SCADA Download Ramp Up Duration
        [25]   // Yeast Cropping FV1-17 SCADA Download Maximum Speed Duration
        [26]   // Yeast Cropping FV1-17 SCADA Download Flush Duration
        [2]   // Yeast Cropping FV1-17 Status
        [2].0   // Yeast Cropping FV1-17 Status Idle
        [2].1   // Yeast Cropping FV1-17 Status Running
        [2].2   // Yeast Cropping FV1-17 Status Held
        [2].3   // Yeast Cropping FV1-17
        [30]   // Yeast Cropping FV1-17 Vessel ID
        [31]   // Yeast Cropping FV1-17 Minimum Speed
        [32]   // Yeast Cropping FV1-17 Maximum Speed
        [33]   // Yeast Cropping FV1-17 Minimum Speed Duration
        [34]   // Yeast Cropping FV1-17 Ramp Up Duration
        [35]   // Yeast Cropping FV1-17 Maximum Speed Duration
        [36]   // Yeast Cropping FV1-17 Flush Duration
        [3]   // Yeast Cropping FV1-17 SCADA Prompts
        [3].0   // Yeast Cropping FV1-17 SCADA Prompts Start
        [3].1   // Yeast Cropping FV1-17 SCADA Prompts Hold
        [3].15   // Yeast Cropping FV1-17 SCADA Prompts Reset
        [3].2   // Yeast Cropping FV1-17 SCADA Prompts Continue
        [3].3   // Yeast Cropping FV1-17 SCADA Prompts Abort
        [3].4   // Yeast Cropping FV1-17 SCADA Prompts Cancel
        [3].5   // Yeast Cropping FV1-17 SCADA Prompts Flush
        [3].6   // Yeast Cropping FV1-17 SCADA Prompts Complete
        [40]   // Yeast Cropping FV1-17 FV File Number
        [41]   // Yeast Cropping FV1-17 Pump Speed
        [42]   // Yeast Cropping FV1-17 Ramp Up Current Time
        [43]   // Yeast Cropping FV1-17
        [4]   // Yeast Cropping FV1-17 SCADA Commands
        [4].0   // Yeast Cropping FV1-17 SCADA Commands Start
        [4].1   // Yeast Cropping FV1-17 SCADA Commands Hold
        [4].2   // Yeast Cropping FV1-17 SCADA Commands Continue
        [4].3   // Yeast Cropping FV1-17 SCADA Commands Abort
        [4].4   // Yeast Cropping FV1-17 SCADA Commands Cancel
        [4].5   // Yeast Cropping FV1-17 SCADA Commands Flush
        [4].6   // Yeast Cropping FV1-17 SCADA Commands Complete
        [50]   // Yeast Cropping FV1-17
        [51]   // Yeast Cropping FV1-17
        [52]   // Yeast Cropping FV1-17
        [53]   // Yeast Cropping FV1-17
        [54]   // Yeast Cropping FV1-17
        [55]   // Yeast Cropping FV1-17
        [56]   // Yeast Cropping FV1-17
        [57]   // Yeast Cropping FV1-17
        [58]   // Yeast Cropping FV1-17 Flush Duration
        [5]   // Yeast Cropping FV1-17 Last SCADA Commands
        [6]   // Yeast Cropping FV1-17 Plant Warning
        [7]   // Yeast Cropping FV1-17 Plant Fault
        [8]   // Yeast Cropping FV1-17 Log Message
        [9]   // Yeast Cropping FV1-17 Plant Item Fault
   FR_N180 : INT[265] := ([100] := 4, [101] := -1, [102] := -1, [103] := -1, [104] := -1, [105] := -1, [106] := -1, [107] := -1, [108] := -1, [109] := -1, [110] := -1, [111] := -1, [112] := -1, [113] := -1, [114] := -1, [115] := -1, [116] := -1, [117] := -1, [118] := -1, [119] := -1, [120] := -1, [121] := -1, [122] := -1, [123] := -1, [124] := -1, [125] := -1, [126] := -1, [127] := -1, [128] := -1, [129] := -1, [130] := -1, [131] := -1, [132] := -1, [133] := -1, [134] := -1, [135] := -1, [136] := -1, [137] := -1, [138] := -1, [139] := -1, [140] := -1, [141] := -1, [142] := -1, [143] := -1, [144] := -1, [145] := -1, [146] := -1, [147] := -1, [148] := -1, [149] := -1);   // Original N File From SLC, No Description Available
        [0]   // Yeast Cropping FV18-25 Step
        [10]   // Yeast Cropping FV18-25 Idle Step Bits
        [10].0   // Yeast Cropping FV18-25 Available
        [10].1   // Yeast Cropping FV18-25 Clean
        [10].2   // Yeast Cropping FV18-25 Command Data Check
        [10].3   // Yeast Cropping FV18-25 Data in Limits Check
        [10].4   // Yeast Cropping FV18-25 FV Vessel Status Check
        [11]   // Yeast Cropping FV18-25 Running Step Bits
        [11].0   // Yeast Cropping FV18-25 Initialise Transfer
        [11].1   // Yeast Cropping FV18-25 Open Route
        [11].2   // Yeast Cropping FV18-25 Minimum Speed
        [11].3   // Yeast Cropping FV18-25 Ramp Up
        [11].4   // Yeast Cropping FV18-25 Maximum Speed
        [11].5   // Yeast Cropping FV18-25 Done
        [11].6   // Yeast Cropping FV18-25 Flush
        [12]   // Yeast Cropping FV18-25 CIP Step Bits
        [12].0   // Yeast Cropping FV18-25 Channel 1 CIP
        [12].1   // Yeast Cropping FV18-25 Channel 1 CIP Complete
        [12].2   // Yeast Cropping FV18-25 Channel 2 CIP
        [12].3   // Yeast Cropping FV18-25 Channel 2 CIP Complete
        [13]   // Yeast Cropping FV18-25 Held Step Bits
        [14].0   // Yeast Cropping FV18-25 Data in Limits Check Vessel Number OK
        [15].0   // Yeast Cropping FV18-25 Auto FV
        [1]   // Yeast Cropping FV18-25 Backup Step
        [20]   // Yeast Cropping FV18-25 SCADA Download Vessel ID
        [21]   // Yeast Cropping FV18-25 SCADA Download Minimum Speed
        [22]   // Yeast Cropping FV18-25 SCADA Download Maximum Speed
        [23]   // Yeast Cropping FV18-25 SCADA Download Minimum Speed Duration
        [24]   // Yeast Cropping FV18-25 SCADA Download Ramp Up Duration
        [25]   // Yeast Cropping FV18-25 SCADA Download Maximum Speed Duration
        [26]   // Yeast Cropping FV18-25 SCADA Download Flush Duration
        [2]   // Yeast Cropping FV18-25 Status
        [2].0   // Yeast Cropping FV18-25 Status Idle
        [2].1   // Yeast Cropping FV18-25 Status Running
        [2].2   // Yeast Cropping FV18-25 Status Held
        [2].3   // Yeast Cropping FV18-25
        [30]   // Yeast Cropping FV18-25 Vessel ID
        [31]   // Yeast Cropping FV18-25 Minimum Speed
        [32]   // Yeast Cropping FV18-25 Maximum Speed
        [33]   // Yeast Cropping FV18-25 Minimum Speed Duration
        [34]   // Yeast Cropping FV18-25 Ramp Up Duration
        [35]   // Yeast Cropping FV18-25 Maximum Speed Duration
        [36]   // Yeast Cropping FV18-25 Flush Duration
        [3]   // Yeast Cropping FV18-25 SCADA Prompts
        [3].0   // Yeast Cropping FV18-25 SCADA Prompts Start
        [3].1   // Yeast Cropping FV18-25 SCADA Prompts Hold
        [3].15   // Yeast Cropping FV18-25 SCADA Prompts Reset
        [3].2   // Yeast Cropping FV18-25 SCADA Prompts Continue
        [3].3   // Yeast Cropping FV18-25 SCADA Prompts Abort
        [3].4   // Yeast Cropping FV18-25 SCADA Prompts Cancel
        [3].5   // Yeast Cropping FV18-25 SCADA Prompts Flush
        [3].6   // Yeast Cropping FV18-25 SCADA Prompts Complete
        [40]   // Yeast Cropping FV18-25 FV File Number
        [41]   // Yeast Cropping FV18-25 Pump Speed
        [42]   // Yeast Cropping FV18-25 Ramp Up Current Time
        [43]   // Yeast Cropping FV18-25
        [4]   // Yeast Cropping FV18-25 SCADA Commands
        [4].0   // Yeast Cropping FV18-25 SCADA Commands Start
        [4].1   // Yeast Cropping FV18-25 SCADA Commands Hold
        [4].2   // Yeast Cropping FV18-25 SCADA Commands Continue
        [4].3   // Yeast Cropping FV18-25 SCADA Commands Abort
        [4].4   // Yeast Cropping FV18-25 SCADA Commands Cancel
        [4].5   // Yeast Cropping FV18-25 SCADA Commands Flush
        [4].6   // Yeast Cropping FV18-25 SCADA Commands Complete
        [50]   // Yeast Cropping FV18-25
        [51]   // Yeast Cropping FV18-25
        [52]   // Yeast Cropping FV18-25
        [53]   // Yeast Cropping FV18-25
        [54]   // Yeast Cropping FV18-25
        [55]   // Yeast Cropping FV18-25
        [56]   // Yeast Cropping FV18-25
        [57]   // Yeast Cropping FV18-25
        [58]   // Yeast Cropping FV18-25 Flush Duration
        [5]   // Yeast Cropping FV18-25 Last SCADA Commands
        [6]   // Yeast Cropping FV18-25 Plant Warning
        [7]   // Yeast Cropping FV18-25 Plant Fault
        [8]   // Yeast Cropping FV18-25 Log Message
        [9]   // Yeast Cropping FV18-25 Plant Item Fault
   FR_N198 : INT[265] := ([0] := -32752);   // Original N File From SLC, No Description Available
   FR_N20 : INT[265] := ([0] := 168, [1] := 50, [2] := 500);   // GENERAL General Purpose Setp oints
        [0]   // Yeast Cropping Timeout
        [2]   // Yeast Cropping Pump CIP Speed
   FR_N200 : INT[265] := ([0] := 2, [2] := 4009, [4] := 4000, [5] := 20000, [7] := 2901, [8] := 5000, [10] := 669, [12] := 8337, [14] := 4000, [15] := 20000, [17] := 2901, [18] := 5000, [20] := 1030, [22] := 3976, [24] := 4000, [25] := 20000, [27] := 2901, [28] := 5000, [30] := 2387, [32] := 10609, [34] := 4000, [35] := 20000, [37] := 2901, [38] := 5000, [40] := 1, [42] := 4001, [44] := 4000, [45] := 20000, [47] := 2901, [48] := 5000, [50] := 1150, [52] := 3994, [54] := 4000, [55] := 20000, [57] := 2901, [58] := 5000, [60] := 6, [62] := 4088, [64] := 4000, [65] := 20000, [67] := 2901, [68] := 5000, [70] := -1, [71] := 2, [72] := 10420, [74] := 4000, [75] := 20000, [77] := 2901, [78] := 5000, [80] := -5, [81] := 2, [82] := 4055, [84] := 4000, [85] := 20000, [87] := 4215, [88] := 5000, [90] := -7, [91] := 2, [92] := 8250, [94] := 4000,
        [95] := 20000, [97] := 4215, [98] := 5000, [100] := -1, [101] := 2, [102] := 3995, [104] := 4000, [105] := 20000, [107] := 4215, [108] := 5000, [110] := 1143, [112] := 8246, [114] := 4000, [115] := 20000, [117] := 4215, [118] := 5000, [120] := -32768, [121] := 2, [124] := 4000, [125] := 20000, [127] := 4000, [130] := -32768, [131] := 2, [134] := 4000, [135] := 20000, [137] := 4000, [140] := -32768, [141] := 2, [144] := 4000, [145] := 20000, [147] := 4000, [150] := -32768, [151] := 2, [154] := 4000, [155] := 20000, [157] := 4000);   // ANALOG_IN Analog Inputs
        [0]   // FV26/PTX01 FV26 top pressure transmitter
        [100]   // FV31/PTX01 FV31 top pressure transmitter
        [101]   // FV31/PTX01 FV31 top pressure Flags
        [101].0   // FV31/PTX01 FV31 top pressure High
        [101].1   // FV31/PTX01 FV31 top pressure Low
        [101].15   // FV31/PTX01 FV31 top pressure Fault
        [102]   // FV31/PTX01 FV31 top pressure mA
        [103]   // FV31/PTX01 FV31 top pressure spare
        [104]   // FV31/PTX01 FV31 top pressure min input
        [105]   // FV31/PTX01 FV31 top pressure max input
        [106]   // FV31/PTX01 FV31 top pressure min scaled
        [107]   // FV31/PTX01 FV31 top pressure max scale
        [108]   // FV31/PTX01 FV31 top pressure High Limit
        [109]   // FV31/PTX01 FV31 top pressure Low Limit
        [10]   // FV26/LTX01 FV26 level transmitter
        [110]   // FV31/LTX01 FV31 level transmitter
        [111]   // FV31/LTX01 FV31 level transmitter Flags
        [111].0   // FV31/LTX01 FV31 level transmitter High
        [111].1   // FV31/LTX01 FV31 level transmitter Low
        [111].15   // FV31/LTX01 FV31 level transmitter Fault
        [112]   // FV31/LTX01 FV31 level transmitter mA
        [113]   // FV31/LTX01 FV31 level transmitter spare
        [114]   // FV31/LTX01 FV31 level transmitter min input
        [115]   // FV31/LTX01 FV31 level transmitter max input
        [116]   // FV31/LTX01 FV31 level transmitter min scaled
        [117]   // FV31/LTX01 FV31 level transmitter max scale
        [118]   // FV31/LTX01 FV31 level transmitter High Limit
        [119]   // FV31/LTX01 FV31 level transmitter Low Limit
        [11]   // FV26/LTX01 FV26 level transmitter Flags
        [11].0   // FV26/LTX01 FV26 level transmitter High
        [11].1   // FV26/LTX01 FV26 level transmitter Low
        [11].15   // FV26/LTX01 FV26 level transmitter Fault
        [121]   // 0 0 0 Flags
        [121].0   // 0 0 0 High
        [121].1   // 0 0 0 Low
        [121].15   // 0 0 0 Fault
        [122]   // 0 0 0 mA
        [123]   // 0 0 0 spare
        [124]   // 0 0 0 min input
        [125]   // 0 0 0 max input
        [126]   // 0 0 0 min scaled
        [127]   // 0 0 0 max scale
        [128]   // 0 0 0 High Limit
        [129]   // 0 0 0 Low Limit
        [12]   // FV26/LTX01 FV26 level transmitter mA
        [131]   // 0 0 0 Flags
        [131].0   // 0 0 0 High
        [131].1   // 0 0 0 Low
        [131].15   // 0 0 0 Fault
        [132]   // 0 0 0 mA
        [133]   // 0 0 0 spare
        [134]   // 0 0 0 min input
        [135]   // 0 0 0 max input
        [136]   // 0 0 0 min scaled
        [137]   // 0 0 0 max scale
        [138]   // 0 0 0 High Limit
        [139]   // 0 0 0 Low Limit
        [13]   // FV26/LTX01 FV26 level transmitter spare
        [141]   // 0 0 0 Flags
        [141].0   // 0 0 0 High
        [141].1   // 0 0 0 Low
        [141].15   // 0 0 0 Fault
        [142]   // 0 0 0 mA
        [143]   // 0 0 0 spare
